(* Logix 5000 project; controller MV vendor 1 type 14 code 217 rev 31.11; software revision 31.00; part 34 of 53 *)
(* tags used below, declared in another part *)
   Alarm_Reset : BOOL;
   Always_Off : BOOL;
   Always_On : BOOL;
   Analog_Fault_No : DINT;
   Analog_Simulation_Enabled : BOOL;
   CLOCK_system_set : BOOL;
   CLOCKsetvalues : DINT[7];
   CWD : CHECKWORD_FLAGS;
   Default_Check_Time : DINT;
   Half_Second_Timer_Off : TIMER;
   Half_Second_Toggle : BOOL;
   MV_B100 : INT[255];   // AT FLAGS
   MV_B3 : INT[255];   // BINARY
   MV_B3_0_1_OUTPUTBIT : BOOL;
   MV_B3_0_2_OUTPUTBIT : BOOL;
   MV_MV10_RTD1_AI : PlantItem;   // MV10_RTD1
   MV_MV10_RTD1_AI_RawInput : ALIAS FOR Remote_IO:2:I.Ch3Data;   // Real Analog Input , Do Not Use In Code
   MV_MV11_RTD1_AI : PlantItem;   // MV11_RTD1
   MV_MV11_RTD1_AI_RawInput : ALIAS FOR Remote_IO:2:I.Ch4Data;   // Real Analog Input , Do Not Use In Code
   MV_MV12_RTD1_AI : PlantItem;   // MV12_RTD1
   MV_MV12_RTD1_AI_RawInput : ALIAS FOR Remote_IO:2:I.Ch5Data;   // Real Analog Input , Do Not Use In Code
   MV_MV13_RTD1_AI : PlantItem;   // MV13_RTD1
   MV_MV13_RTD1_AI_RawInput : ALIAS FOR Remote_IO:3:I.Ch0Data;   // Real Analog Input , Do Not Use In Code
   MV_MV14_RTD1_AI : PlantItem;   // MV14_RTD1
   MV_MV14_RTD1_AI_RawInput : ALIAS FOR Remote_IO:3:I.Ch1Data;   // Real Analog Input , Do Not Use In Code
   MV_MV15_RTD1_AI : PlantItem;   // MV15_RTD1
   MV_MV15_RTD1_AI_RawInput : ALIAS FOR Remote_IO:3:I.Ch2Data;   // Real Analog Input , Do Not Use In Code
   MV_MV16_RTD1_AI : PlantItem;   // MV16_RTD1
   MV_MV16_RTD1_AI_RawInput : ALIAS FOR Remote_IO:3:I.Ch3Data;   // Real Analog Input , Do Not Use In Code
   MV_MV17_RTD1_AI : PlantItem;   // MV17_RTD1
   MV_MV17_RTD1_AI_RawInput : ALIAS FOR Remote_IO:3:I.Ch4Data;   // Real Analog Input , Do Not Use In Code
   MV_MV1_RTD1_AI : PlantItem;   // MV1_RTD1
   MV_MV1_RTD1_AI_RawInput : ALIAS FOR Remote_IO:1:I.Ch0Data;   // Real Analog Input , Do Not Use In Code
   MV_MV2_RTD1_AI : PlantItem;   // MV2_RTD1
   MV_MV2_RTD1_AI_RawInput : ALIAS FOR Remote_IO:1:I.Ch1Data;   // Real Analog Input , Do Not Use In Code
   MV_MV3_RTD1_AI : PlantItem;   // MV3_RTD1
   MV_MV3_RTD1_AI_RawInput : ALIAS FOR Remote_IO:1:I.Ch2Data;   // Real Analog Input , Do Not Use In Code
   MV_MV4_RTD1_AI : PlantItem;   // MV4_RTD1
   MV_MV4_RTD1_AI_RawInput : ALIAS FOR Remote_IO:1:I.Ch3Data;   // Real Analog Input , Do Not Use In Code
   MV_MV5_RTD1_AI : PlantItem;   // MV5_RTD1
   MV_MV5_RTD1_AI_RawInput : ALIAS FOR Remote_IO:1:I.Ch4Data;   // Real Analog Input , Do Not Use In Code
   MV_MV6_RTD1_AI : PlantItem;   // MV6_RTD1
   MV_MV6_RTD1_AI_RawInput : ALIAS FOR Remote_IO:1:I.Ch5Data;   // Real Analog Input , Do Not Use In Code
   MV_MV7_RTD1_AI : PlantItem;   // MV7_RTD1
   MV_MV7_RTD1_AI_RawInput : ALIAS FOR Remote_IO:2:I.Ch0Data;   // Real Analog Input , Do Not Use In Code
   MV_MV8_RTD1_AI : PlantItem;   // MV8_RTD1
   MV_MV8_RTD1_AI_RawInput : ALIAS FOR Remote_IO:2:I.Ch1Data;   // Real Analog Input , Do Not Use In Code
   MV_MV9_RTD1_AI : PlantItem;   // MV9_RTD1
   MV_MV9_RTD1_AI_RawInput : ALIAS FOR Remote_IO:2:I.Ch2Data;   // Real Analog Input , Do Not Use In Code
   MV_N12 : INT[255];   // SYS_PARMS System Parameter Fil e
   MV_SFile : INT[255];   // SLC Equivalent System File, So Original Code Can Remain
   MV_T4 : TIMER[20];
   One_Minute_One_Scan : BOOL;
   One_Minute_One_Scan_Timer : TIMER;
   One_sec_toggle : DINT;
   One_Second_1_scan : BOOL;
   One_Second_One_Scan : ALIAS FOR One_Second_1_scan;
   One_Second_Toggle : BOOL;
   One_Second_Toggle_Valid_Groups : BOOL;
   overrange_RIO_analog_value : REAL;
   scada_watchdog : DINT;
   underrange_RIO_analog_value : REAL;
(* MV_Common, continued *)

ROUTINE general_timers   (* ladder *)
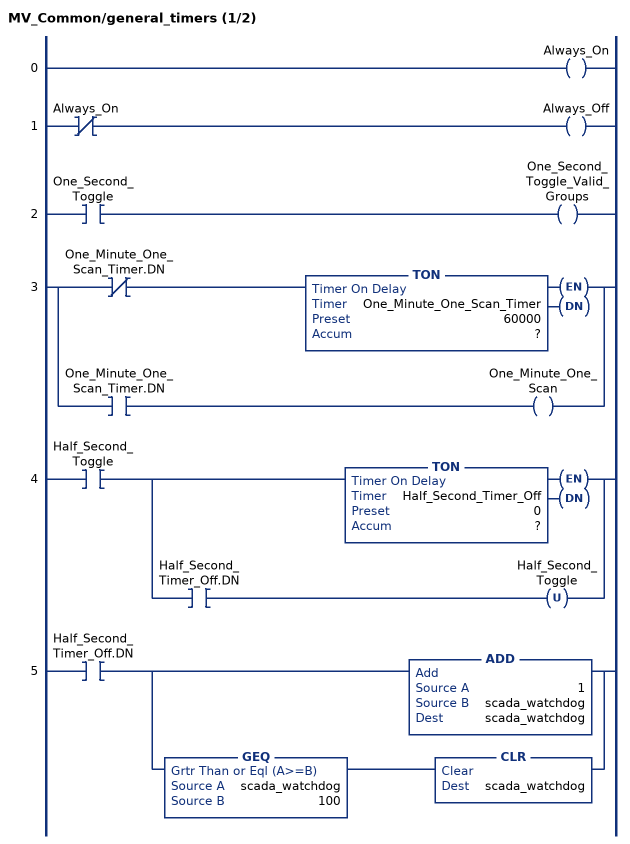
   0: OTE(Always_On);
   1: XIO(Always_On)OTE(Always_Off);
   2: XIC(One_Second_Toggle)OTE(One_Second_Toggle_Valid_Groups);
   3: [XIO(One_Minute_One_Scan_Timer.DN) TON(One_Minute_One_Scan_Timer,?,?) ,XIC(One_Minute_One_Scan_Timer.DN) OTE(One_Minute_One_Scan) ];
   4: XIC(Half_Second_Toggle)[TON(Half_Second_Timer_Off,?,?) ,XIC(Half_Second_Timer_Off.DN) OTU(Half_Second_Toggle) ];
   5: XIC(Half_Second_Timer_Off.DN)[ADD(1,scada_watchdog,scada_watchdog) ,GEQ(scada_watchdog,100) CLR(scada_watchdog) ];
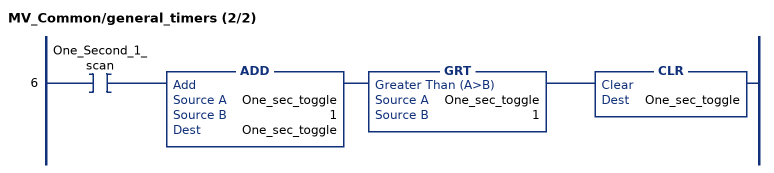
   6: XIC(One_Second_1_scan)ADD(One_sec_toggle,1,One_sec_toggle)GRT(One_sec_toggle,1)CLR(One_sec_toggle);
END_ROUTINE

ROUTINE MainRoutine   (* ladder *)
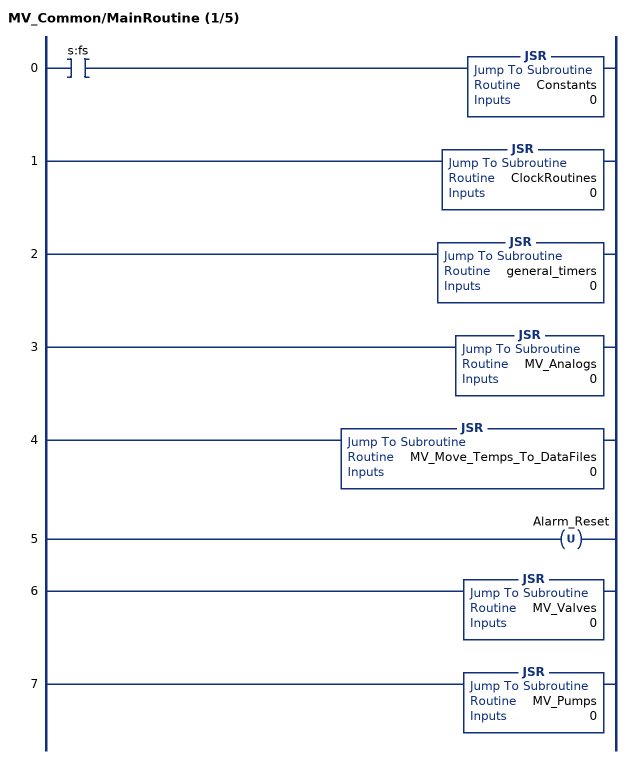
   0: XIC(s:fs)JSR(Constants,0);
   1: JSR(ClockRoutines,0);
   2: JSR(general_timers,0);
   3: JSR(MV_Analogs,0);
   4: JSR(MV_Move_Temps_To_DataFiles,0);
   5: OTU(Alarm_Reset);
   6: JSR(MV_Valves,0);
   7: JSR(MV_Pumps,0);
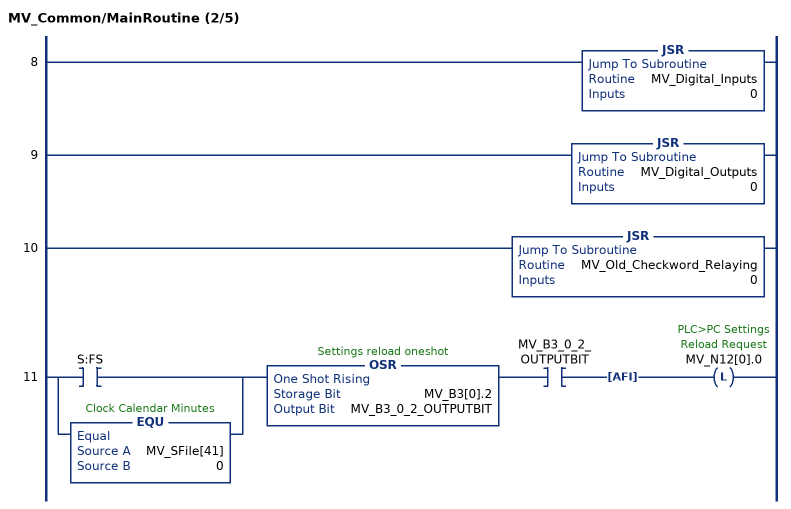
   8: JSR(MV_Digital_Inputs,0);
   9: JSR(MV_Digital_Outputs,0);
   10: JSR(MV_Old_Checkword_Relaying,0);
   11: [XIC(S:FS) ,EQU(MV_SFile[41],0) ]OSR(MV_B3[0].2,MV_B3_0_2_OUTPUTBIT)XIC(MV_B3_0_2_OUTPUTBIT)AFI()OTL(MV_N12[0].0);
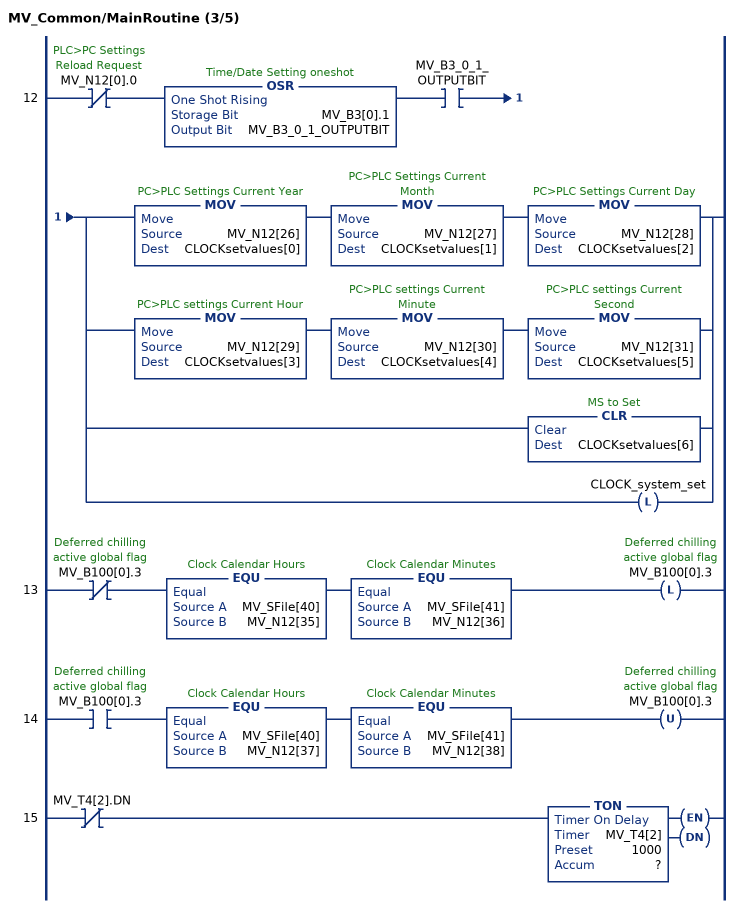
   12: XIO(MV_N12[0].0)OSR(MV_B3[0].1,MV_B3_0_1_OUTPUTBIT)XIC(MV_B3_0_1_OUTPUTBIT)[MOV(MV_N12[26],CLOCKsetvalues[0]) MOV(MV_N12[27],CLOCKsetvalues[1]) MOV(MV_N12[28],CLOCKsetvalues[2]) ,MOV(MV_N12[29],CLOCKsetvalues[3]) MOV(MV_N12[30],CLOCKsetvalues[4]) MOV(MV_N12[31],CLOCKsetvalues[5]) ,CLR(CLOCKsetvalues[6]) ,OTL(CLOCK_system_set) ];
   13: XIO(MV_B100[0].3)EQU(MV_SFile[40],MV_N12[35])EQU(MV_SFile[41],MV_N12[36])OTL(MV_B100[0].3);
   14: XIC(MV_B100[0].3)EQU(MV_SFile[40],MV_N12[37])EQU(MV_SFile[41],MV_N12[38])OTU(MV_B100[0].3);
   15: XIO(MV_T4[2].DN)TON(MV_T4[2],?,?);
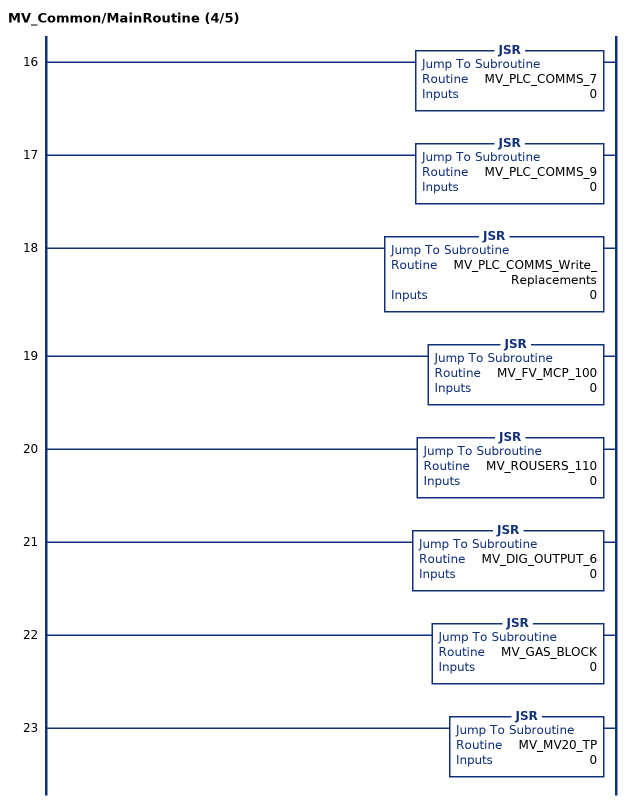
   16: JSR(MV_PLC_COMMS_7,0);
   17: JSR(MV_PLC_COMMS_9,0);
   18: JSR(MV_PLC_COMMS_Write_Replacements,0);
   19: JSR(MV_FV_MCP_100,0);
   20: JSR(MV_ROUSERS_110,0);
   21: JSR(MV_DIG_OUTPUT_6,0);
   22: JSR(MV_GAS_BLOCK,0);
   23: JSR(MV_MV20_TP,0);
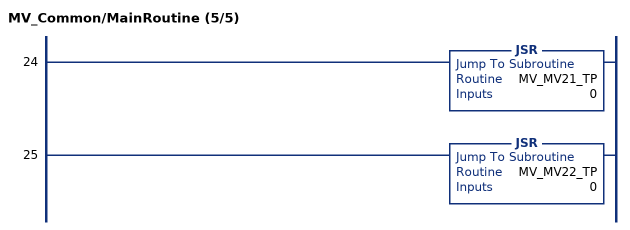
   24: JSR(MV_MV21_TP,0);
   25: JSR(MV_MV22_TP,0);
END_ROUTINE

ROUTINE MV_Analogs   (* ladder *)
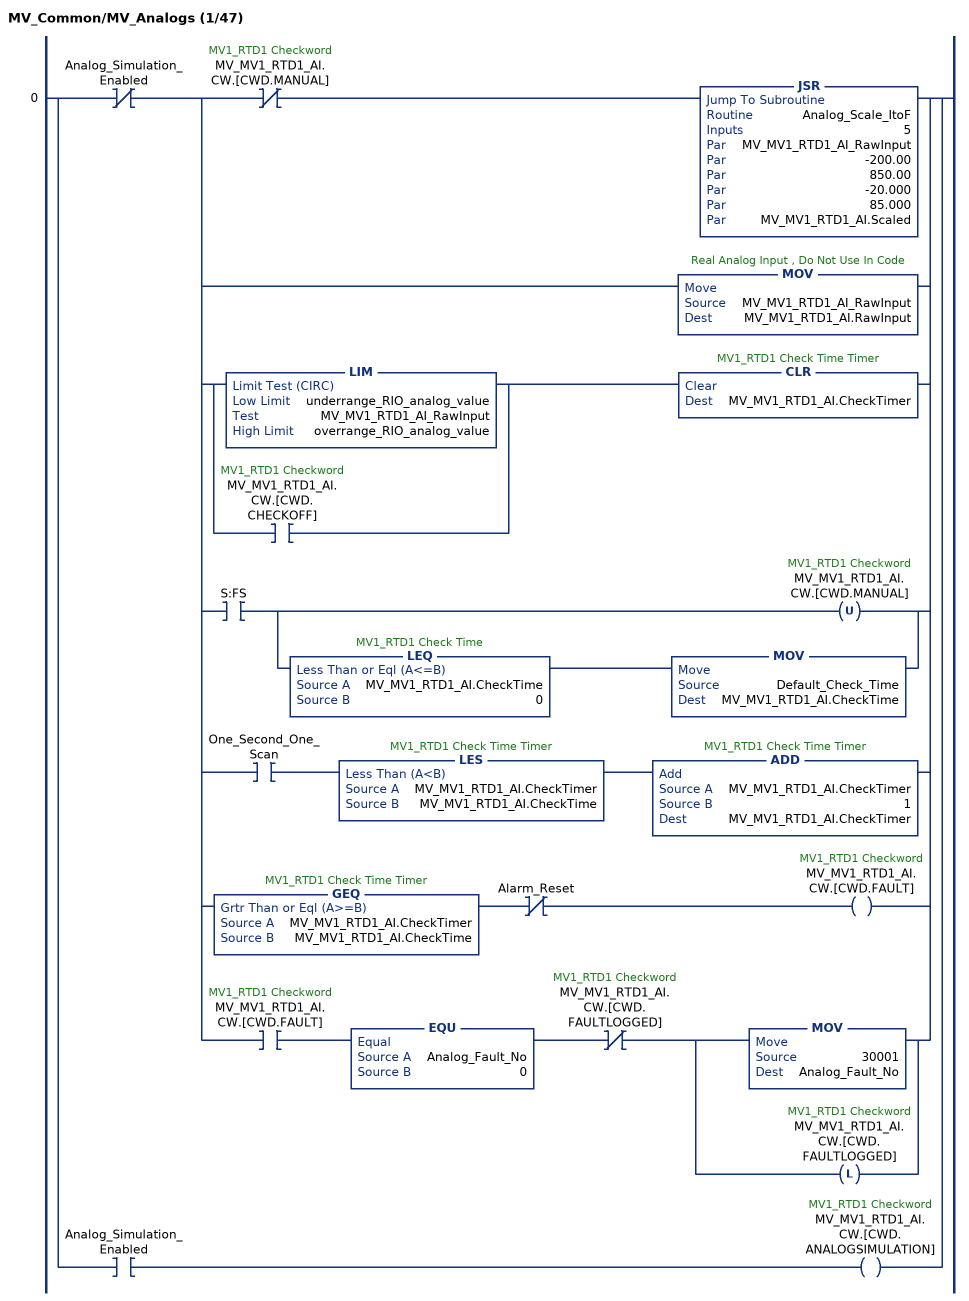
   0: [XIO(Analog_Simulation_Enabled) [XIO(MV_MV1_RTD1_AI.CW.[CWD.MANUAL]) JSR(Analog_Scale_ItoF,5,MV_MV1_RTD1_AI_RawInput,-200.00,850.00,-20.000,85.000,MV_MV1_RTD1_AI.Scaled) ,MOV(MV_MV1_RTD1_AI_RawInput,MV_MV1_RTD1_AI.RawInput) ,[LIM(underrange_RIO_analog_value,MV_MV1_RTD1_AI_RawInput,overrange_RIO_analog_value) ,XIC(MV_MV1_RTD1_AI.CW.[CWD.CHECKOFF]) ] CLR(MV_MV1_RTD1_AI.CheckTimer) ,XIC(S:FS) [OTU(MV_MV1_RTD1_AI.CW.[CWD.MANUAL]) ,LEQ(MV_MV1_RTD1_AI.CheckTime,0) MOV(Default_Check_Time,MV_MV1_RTD1_AI.CheckTime) ] ,XIC(One_Second_One_Scan) LES(MV_MV1_RTD1_AI.CheckTimer,MV_MV1_RTD1_AI.CheckTime) ADD(MV_MV1_RTD1_AI.CheckTimer,1,MV_MV1_RTD1_AI.CheckTimer) ,GEQ(MV_MV1_RTD1_AI.CheckTimer,MV_MV1_RTD1_AI.CheckTime) XIO(Alarm_Reset) OTE(MV_MV1_RTD1_AI.CW.[CWD.FAULT]) ,XIC(MV_MV1_RTD1_AI.CW.[CWD.FAULT]) EQU(Analog_Fault_No,0) XIO(MV_MV1_RTD1_AI.CW.[CWD.FAULTLOGGED]) [MOV(30001,Analog_Fault_No) ,OTL(MV_MV1_RTD1_AI.CW.[CWD.FAULTLOGGED]) ] ] ,XIC(Analog_Simulation_Enabled) OTE(MV_MV1_RTD1_AI.CW.[CWD.ANALOGSIMULATION]) ];
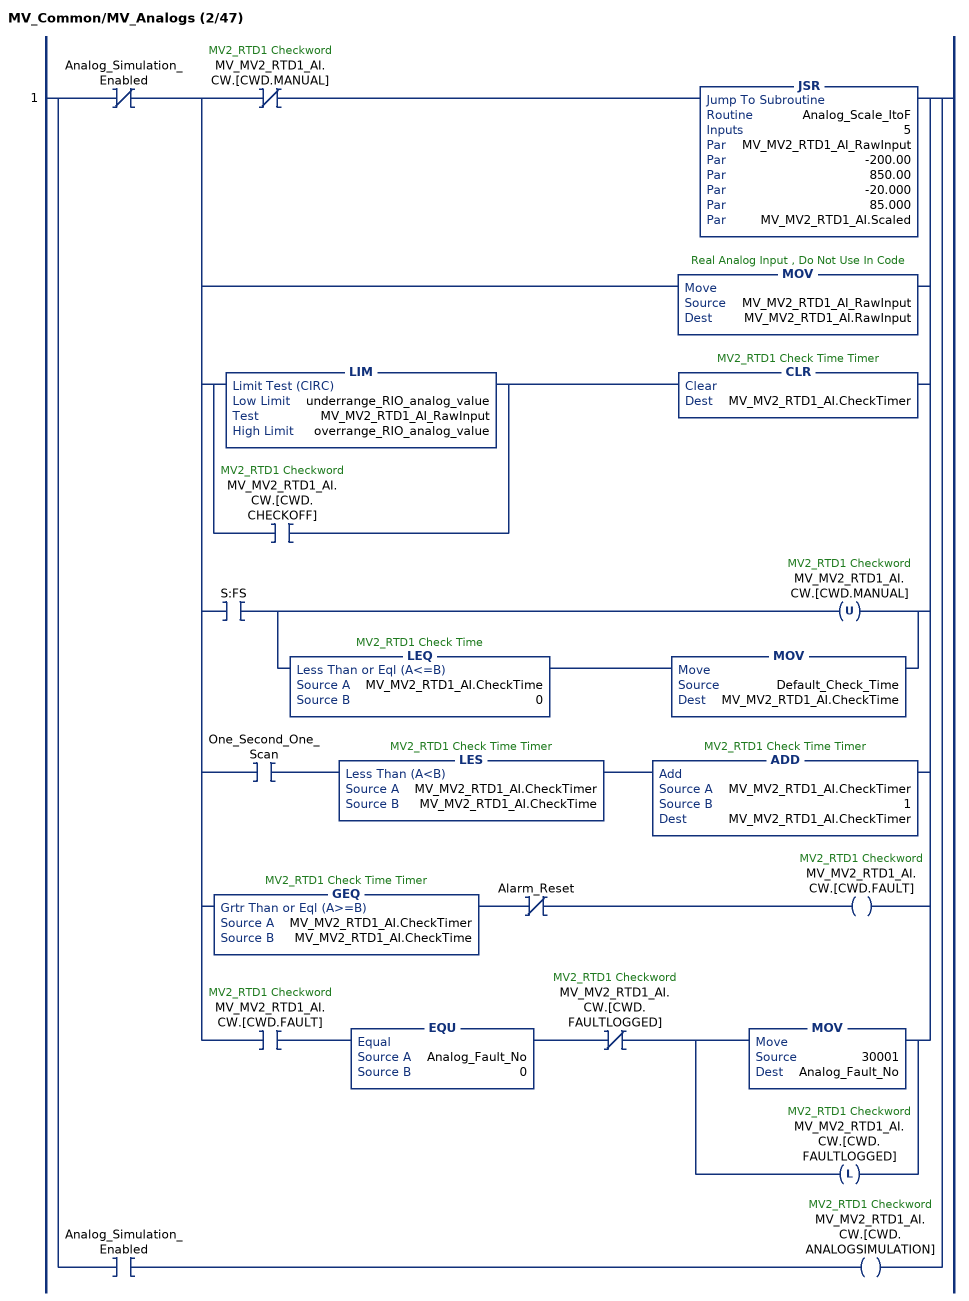
   1: [XIO(Analog_Simulation_Enabled) [XIO(MV_MV2_RTD1_AI.CW.[CWD.MANUAL]) JSR(Analog_Scale_ItoF,5,MV_MV2_RTD1_AI_RawInput,-200.00,850.00,-20.000,85.000,MV_MV2_RTD1_AI.Scaled) ,MOV(MV_MV2_RTD1_AI_RawInput,MV_MV2_RTD1_AI.RawInput) ,[LIM(underrange_RIO_analog_value,MV_MV2_RTD1_AI_RawInput,overrange_RIO_analog_value) ,XIC(MV_MV2_RTD1_AI.CW.[CWD.CHECKOFF]) ] CLR(MV_MV2_RTD1_AI.CheckTimer) ,XIC(S:FS) [OTU(MV_MV2_RTD1_AI.CW.[CWD.MANUAL]) ,LEQ(MV_MV2_RTD1_AI.CheckTime,0) MOV(Default_Check_Time,MV_MV2_RTD1_AI.CheckTime) ] ,XIC(One_Second_One_Scan) LES(MV_MV2_RTD1_AI.CheckTimer,MV_MV2_RTD1_AI.CheckTime) ADD(MV_MV2_RTD1_AI.CheckTimer,1,MV_MV2_RTD1_AI.CheckTimer) ,GEQ(MV_MV2_RTD1_AI.CheckTimer,MV_MV2_RTD1_AI.CheckTime) XIO(Alarm_Reset) OTE(MV_MV2_RTD1_AI.CW.[CWD.FAULT]) ,XIC(MV_MV2_RTD1_AI.CW.[CWD.FAULT]) EQU(Analog_Fault_No,0) XIO(MV_MV2_RTD1_AI.CW.[CWD.FAULTLOGGED]) [MOV(30001,Analog_Fault_No) ,OTL(MV_MV2_RTD1_AI.CW.[CWD.FAULTLOGGED]) ] ] ,XIC(Analog_Simulation_Enabled) OTE(MV_MV2_RTD1_AI.CW.[CWD.ANALOGSIMULATION]) ];
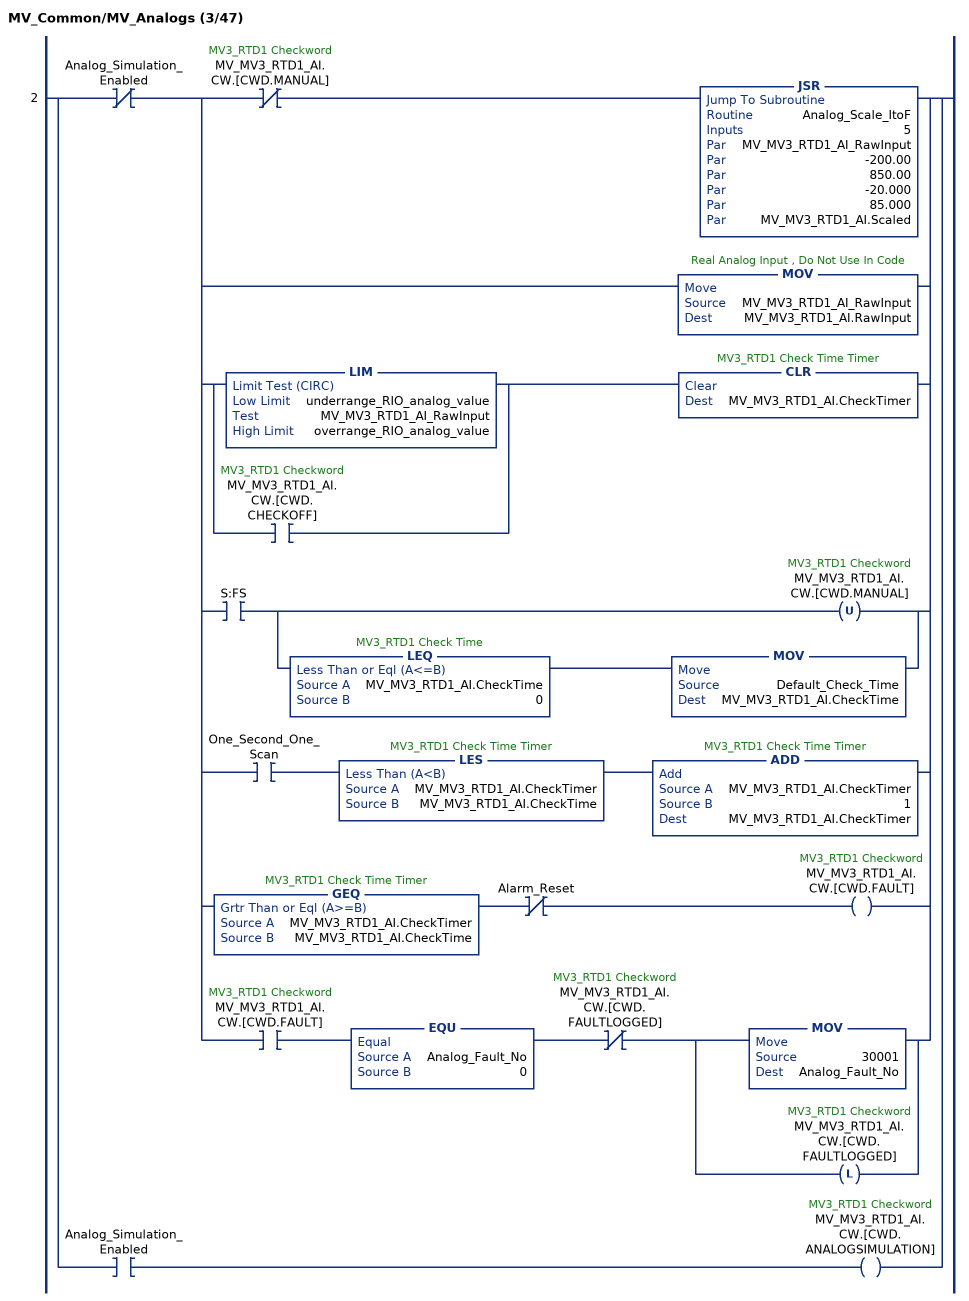
   2: [XIO(Analog_Simulation_Enabled) [XIO(MV_MV3_RTD1_AI.CW.[CWD.MANUAL]) JSR(Analog_Scale_ItoF,5,MV_MV3_RTD1_AI_RawInput,-200.00,850.00,-20.000,85.000,MV_MV3_RTD1_AI.Scaled) ,MOV(MV_MV3_RTD1_AI_RawInput,MV_MV3_RTD1_AI.RawInput) ,[LIM(underrange_RIO_analog_value,MV_MV3_RTD1_AI_RawInput,overrange_RIO_analog_value) ,XIC(MV_MV3_RTD1_AI.CW.[CWD.CHECKOFF]) ] CLR(MV_MV3_RTD1_AI.CheckTimer) ,XIC(S:FS) [OTU(MV_MV3_RTD1_AI.CW.[CWD.MANUAL]) ,LEQ(MV_MV3_RTD1_AI.CheckTime,0) MOV(Default_Check_Time,MV_MV3_RTD1_AI.CheckTime) ] ,XIC(One_Second_One_Scan) LES(MV_MV3_RTD1_AI.CheckTimer,MV_MV3_RTD1_AI.CheckTime) ADD(MV_MV3_RTD1_AI.CheckTimer,1,MV_MV3_RTD1_AI.CheckTimer) ,GEQ(MV_MV3_RTD1_AI.CheckTimer,MV_MV3_RTD1_AI.CheckTime) XIO(Alarm_Reset) OTE(MV_MV3_RTD1_AI.CW.[CWD.FAULT]) ,XIC(MV_MV3_RTD1_AI.CW.[CWD.FAULT]) EQU(Analog_Fault_No,0) XIO(MV_MV3_RTD1_AI.CW.[CWD.FAULTLOGGED]) [MOV(30001,Analog_Fault_No) ,OTL(MV_MV3_RTD1_AI.CW.[CWD.FAULTLOGGED]) ] ] ,XIC(Analog_Simulation_Enabled) OTE(MV_MV3_RTD1_AI.CW.[CWD.ANALOGSIMULATION]) ];
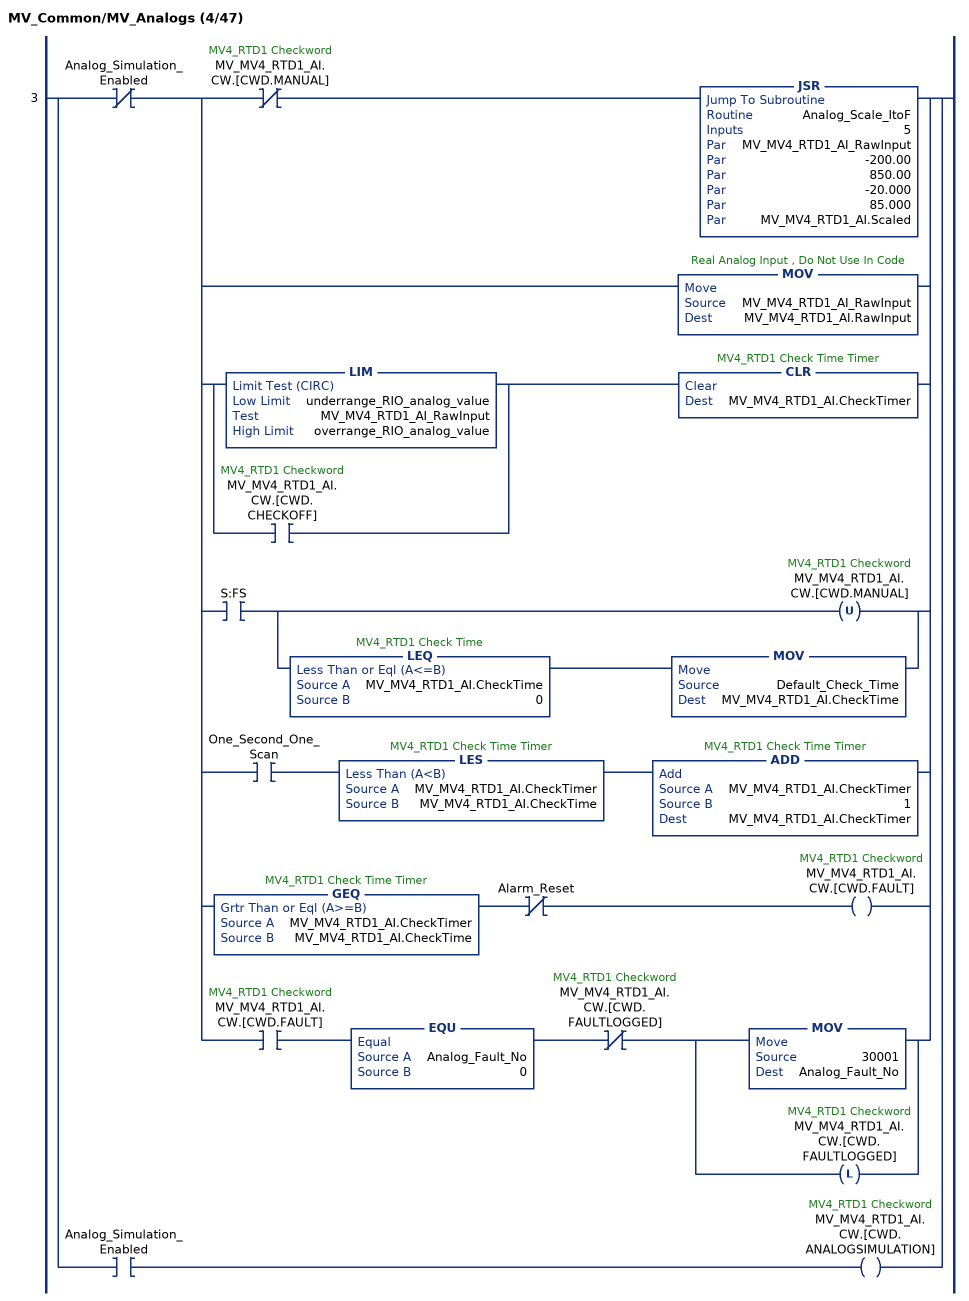
   3: [XIO(Analog_Simulation_Enabled) [XIO(MV_MV4_RTD1_AI.CW.[CWD.MANUAL]) JSR(Analog_Scale_ItoF,5,MV_MV4_RTD1_AI_RawInput,-200.00,850.00,-20.000,85.000,MV_MV4_RTD1_AI.Scaled) ,MOV(MV_MV4_RTD1_AI_RawInput,MV_MV4_RTD1_AI.RawInput) ,[LIM(underrange_RIO_analog_value,MV_MV4_RTD1_AI_RawInput,overrange_RIO_analog_value) ,XIC(MV_MV4_RTD1_AI.CW.[CWD.CHECKOFF]) ] CLR(MV_MV4_RTD1_AI.CheckTimer) ,XIC(S:FS) [OTU(MV_MV4_RTD1_AI.CW.[CWD.MANUAL]) ,LEQ(MV_MV4_RTD1_AI.CheckTime,0) MOV(Default_Check_Time,MV_MV4_RTD1_AI.CheckTime) ] ,XIC(One_Second_One_Scan) LES(MV_MV4_RTD1_AI.CheckTimer,MV_MV4_RTD1_AI.CheckTime) ADD(MV_MV4_RTD1_AI.CheckTimer,1,MV_MV4_RTD1_AI.CheckTimer) ,GEQ(MV_MV4_RTD1_AI.CheckTimer,MV_MV4_RTD1_AI.CheckTime) XIO(Alarm_Reset) OTE(MV_MV4_RTD1_AI.CW.[CWD.FAULT]) ,XIC(MV_MV4_RTD1_AI.CW.[CWD.FAULT]) EQU(Analog_Fault_No,0) XIO(MV_MV4_RTD1_AI.CW.[CWD.FAULTLOGGED]) [MOV(30001,Analog_Fault_No) ,OTL(MV_MV4_RTD1_AI.CW.[CWD.FAULTLOGGED]) ] ] ,XIC(Analog_Simulation_Enabled) OTE(MV_MV4_RTD1_AI.CW.[CWD.ANALOGSIMULATION]) ];
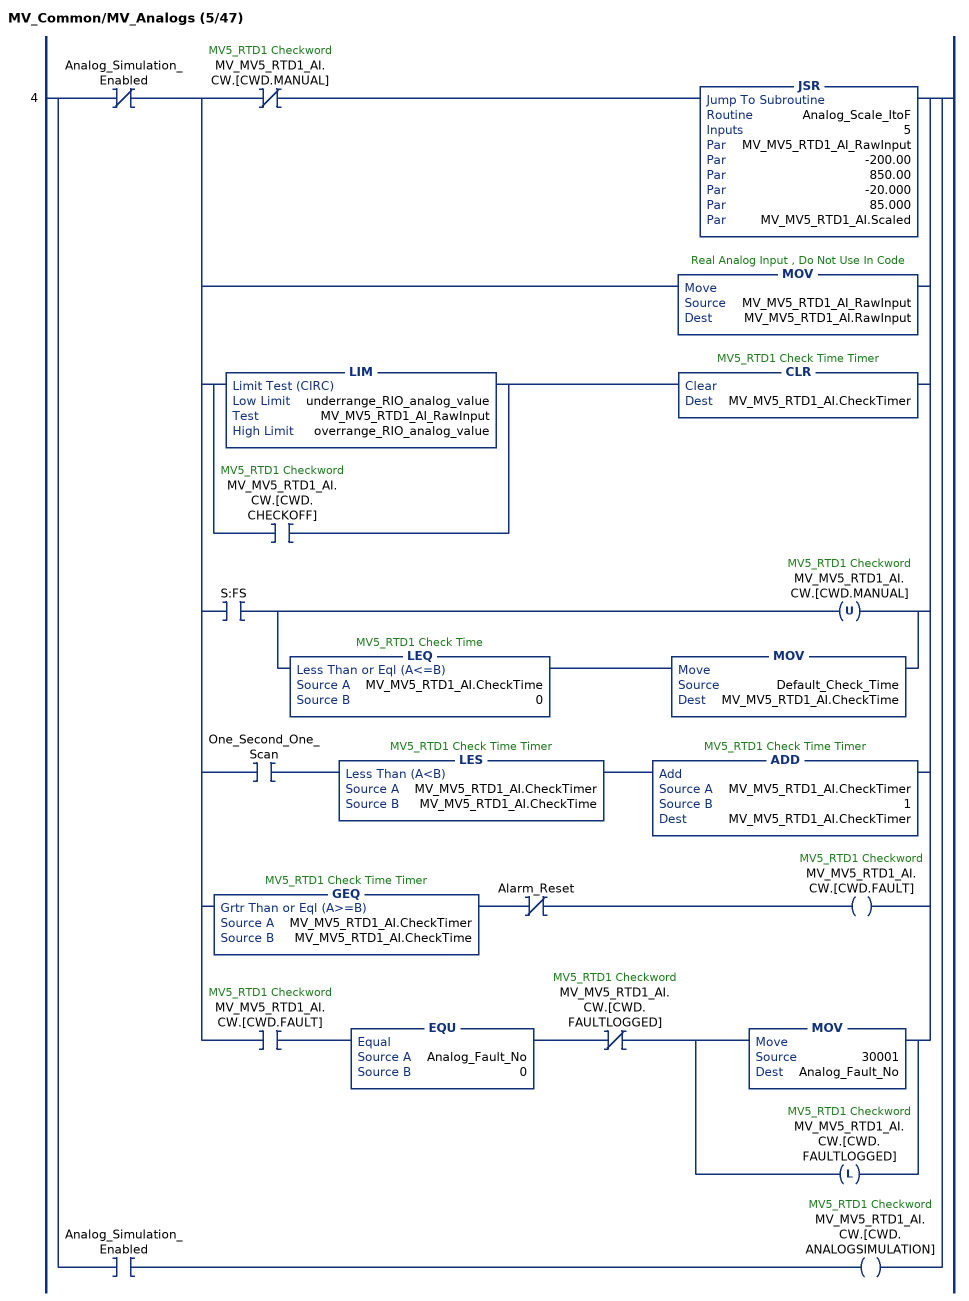
   4: [XIO(Analog_Simulation_Enabled) [XIO(MV_MV5_RTD1_AI.CW.[CWD.MANUAL]) JSR(Analog_Scale_ItoF,5,MV_MV5_RTD1_AI_RawInput,-200.00,850.00,-20.000,85.000,MV_MV5_RTD1_AI.Scaled) ,MOV(MV_MV5_RTD1_AI_RawInput,MV_MV5_RTD1_AI.RawInput) ,[LIM(underrange_RIO_analog_value,MV_MV5_RTD1_AI_RawInput,overrange_RIO_analog_value) ,XIC(MV_MV5_RTD1_AI.CW.[CWD.CHECKOFF]) ] CLR(MV_MV5_RTD1_AI.CheckTimer) ,XIC(S:FS) [OTU(MV_MV5_RTD1_AI.CW.[CWD.MANUAL]) ,LEQ(MV_MV5_RTD1_AI.CheckTime,0) MOV(Default_Check_Time,MV_MV5_RTD1_AI.CheckTime) ] ,XIC(One_Second_One_Scan) LES(MV_MV5_RTD1_AI.CheckTimer,MV_MV5_RTD1_AI.CheckTime) ADD(MV_MV5_RTD1_AI.CheckTimer,1,MV_MV5_RTD1_AI.CheckTimer) ,GEQ(MV_MV5_RTD1_AI.CheckTimer,MV_MV5_RTD1_AI.CheckTime) XIO(Alarm_Reset) OTE(MV_MV5_RTD1_AI.CW.[CWD.FAULT]) ,XIC(MV_MV5_RTD1_AI.CW.[CWD.FAULT]) EQU(Analog_Fault_No,0) XIO(MV_MV5_RTD1_AI.CW.[CWD.FAULTLOGGED]) [MOV(30001,Analog_Fault_No) ,OTL(MV_MV5_RTD1_AI.CW.[CWD.FAULTLOGGED]) ] ] ,XIC(Analog_Simulation_Enabled) OTE(MV_MV5_RTD1_AI.CW.[CWD.ANALOGSIMULATION]) ];
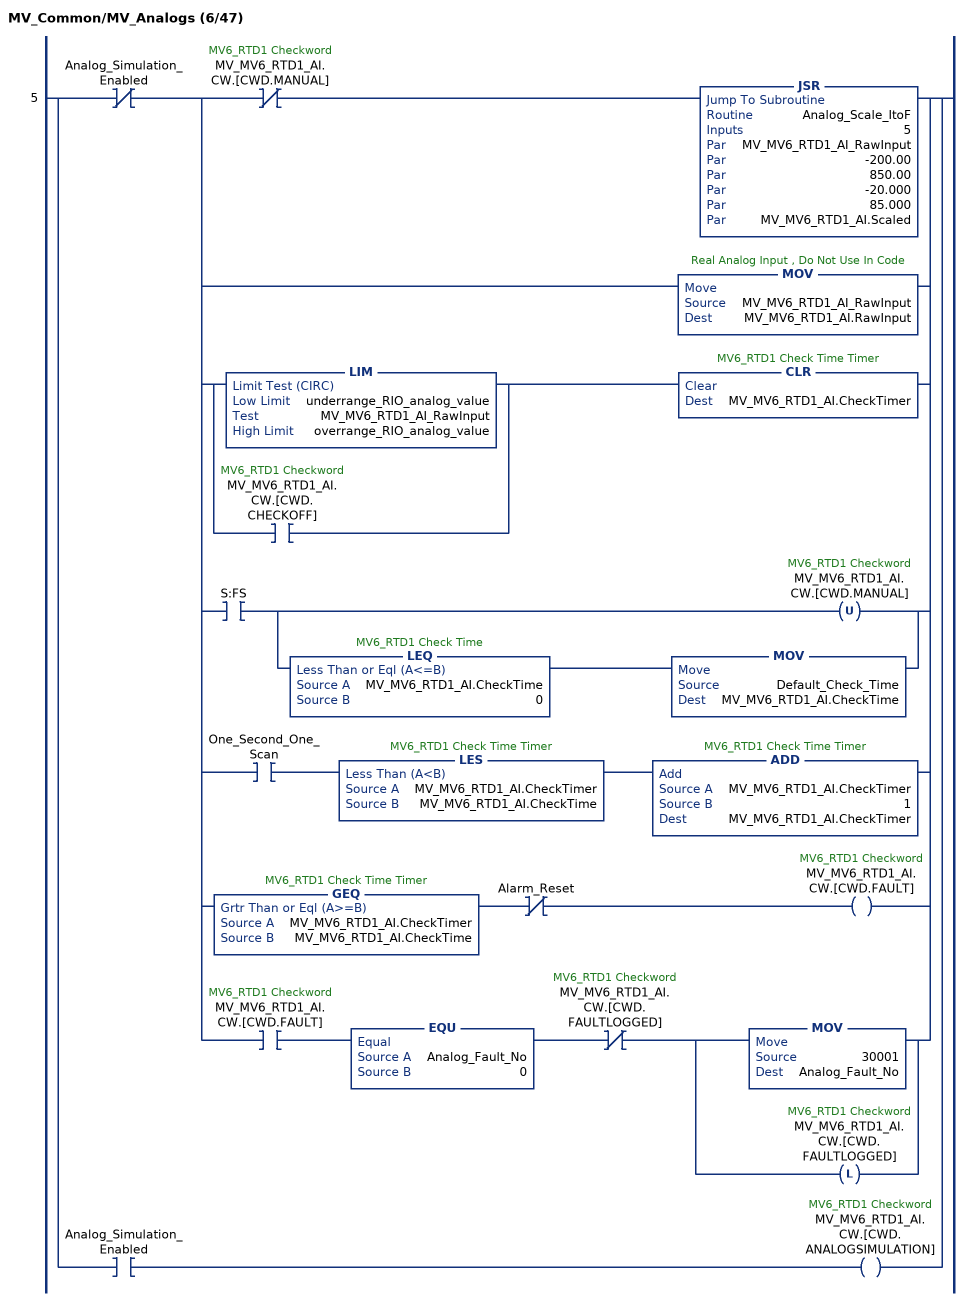
   5: [XIO(Analog_Simulation_Enabled) [XIO(MV_MV6_RTD1_AI.CW.[CWD.MANUAL]) JSR(Analog_Scale_ItoF,5,MV_MV6_RTD1_AI_RawInput,-200.00,850.00,-20.000,85.000,MV_MV6_RTD1_AI.Scaled) ,MOV(MV_MV6_RTD1_AI_RawInput,MV_MV6_RTD1_AI.RawInput) ,[LIM(underrange_RIO_analog_value,MV_MV6_RTD1_AI_RawInput,overrange_RIO_analog_value) ,XIC(MV_MV6_RTD1_AI.CW.[CWD.CHECKOFF]) ] CLR(MV_MV6_RTD1_AI.CheckTimer) ,XIC(S:FS) [OTU(MV_MV6_RTD1_AI.CW.[CWD.MANUAL]) ,LEQ(MV_MV6_RTD1_AI.CheckTime,0) MOV(Default_Check_Time,MV_MV6_RTD1_AI.CheckTime) ] ,XIC(One_Second_One_Scan) LES(MV_MV6_RTD1_AI.CheckTimer,MV_MV6_RTD1_AI.CheckTime) ADD(MV_MV6_RTD1_AI.CheckTimer,1,MV_MV6_RTD1_AI.CheckTimer) ,GEQ(MV_MV6_RTD1_AI.CheckTimer,MV_MV6_RTD1_AI.CheckTime) XIO(Alarm_Reset) OTE(MV_MV6_RTD1_AI.CW.[CWD.FAULT]) ,XIC(MV_MV6_RTD1_AI.CW.[CWD.FAULT]) EQU(Analog_Fault_No,0) XIO(MV_MV6_RTD1_AI.CW.[CWD.FAULTLOGGED]) [MOV(30001,Analog_Fault_No) ,OTL(MV_MV6_RTD1_AI.CW.[CWD.FAULTLOGGED]) ] ] ,XIC(Analog_Simulation_Enabled) OTE(MV_MV6_RTD1_AI.CW.[CWD.ANALOGSIMULATION]) ];
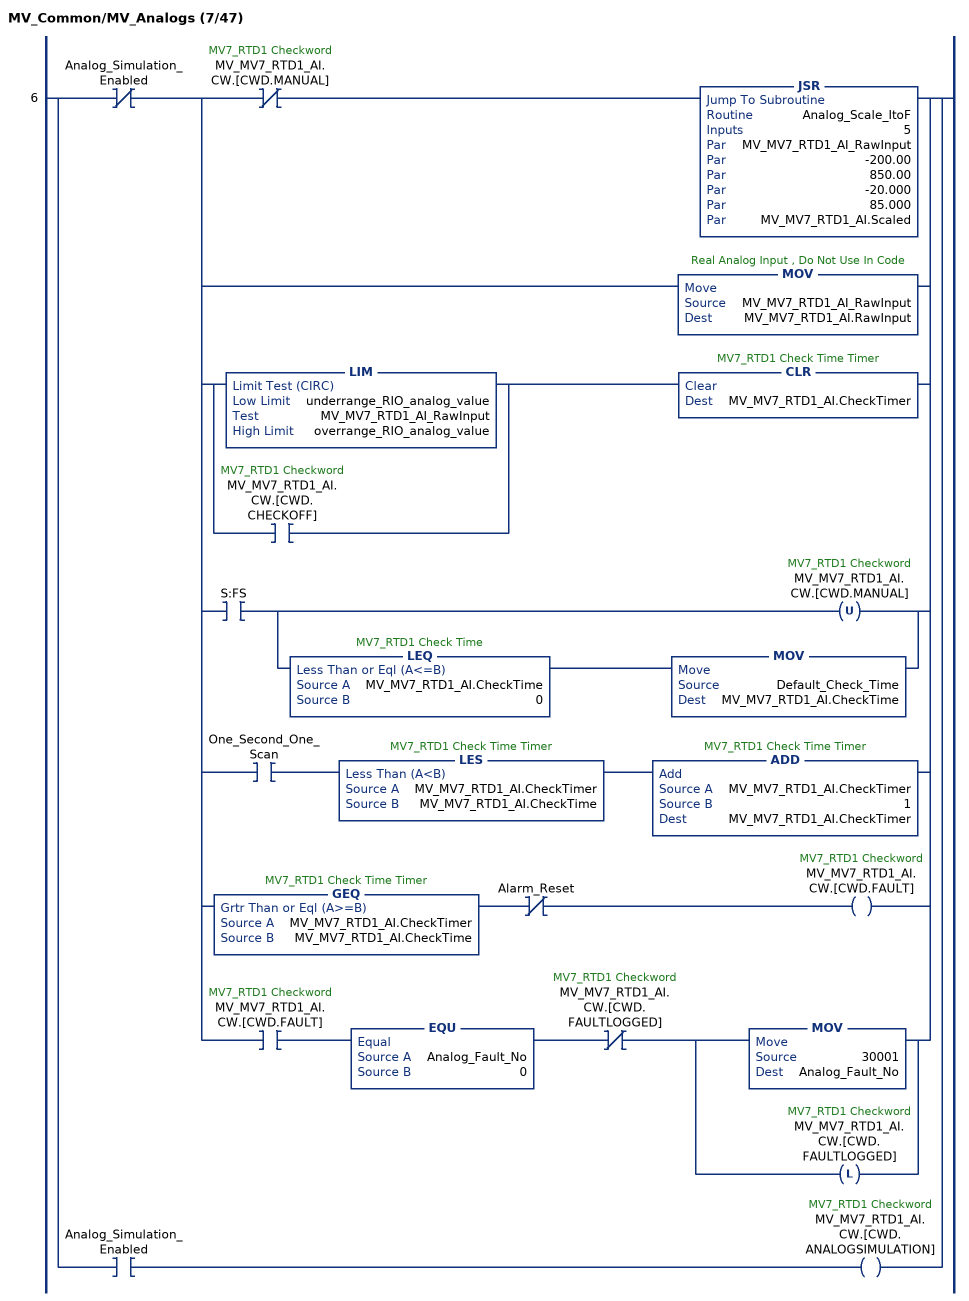
   6: [XIO(Analog_Simulation_Enabled) [XIO(MV_MV7_RTD1_AI.CW.[CWD.MANUAL]) JSR(Analog_Scale_ItoF,5,MV_MV7_RTD1_AI_RawInput,-200.00,850.00,-20.000,85.000,MV_MV7_RTD1_AI.Scaled) ,MOV(MV_MV7_RTD1_AI_RawInput,MV_MV7_RTD1_AI.RawInput) ,[LIM(underrange_RIO_analog_value,MV_MV7_RTD1_AI_RawInput,overrange_RIO_analog_value) ,XIC(MV_MV7_RTD1_AI.CW.[CWD.CHECKOFF]) ] CLR(MV_MV7_RTD1_AI.CheckTimer) ,XIC(S:FS) [OTU(MV_MV7_RTD1_AI.CW.[CWD.MANUAL]) ,LEQ(MV_MV7_RTD1_AI.CheckTime,0) MOV(Default_Check_Time,MV_MV7_RTD1_AI.CheckTime) ] ,XIC(One_Second_One_Scan) LES(MV_MV7_RTD1_AI.CheckTimer,MV_MV7_RTD1_AI.CheckTime) ADD(MV_MV7_RTD1_AI.CheckTimer,1,MV_MV7_RTD1_AI.CheckTimer) ,GEQ(MV_MV7_RTD1_AI.CheckTimer,MV_MV7_RTD1_AI.CheckTime) XIO(Alarm_Reset) OTE(MV_MV7_RTD1_AI.CW.[CWD.FAULT]) ,XIC(MV_MV7_RTD1_AI.CW.[CWD.FAULT]) EQU(Analog_Fault_No,0) XIO(MV_MV7_RTD1_AI.CW.[CWD.FAULTLOGGED]) [MOV(30001,Analog_Fault_No) ,OTL(MV_MV7_RTD1_AI.CW.[CWD.FAULTLOGGED]) ] ] ,XIC(Analog_Simulation_Enabled) OTE(MV_MV7_RTD1_AI.CW.[CWD.ANALOGSIMULATION]) ];